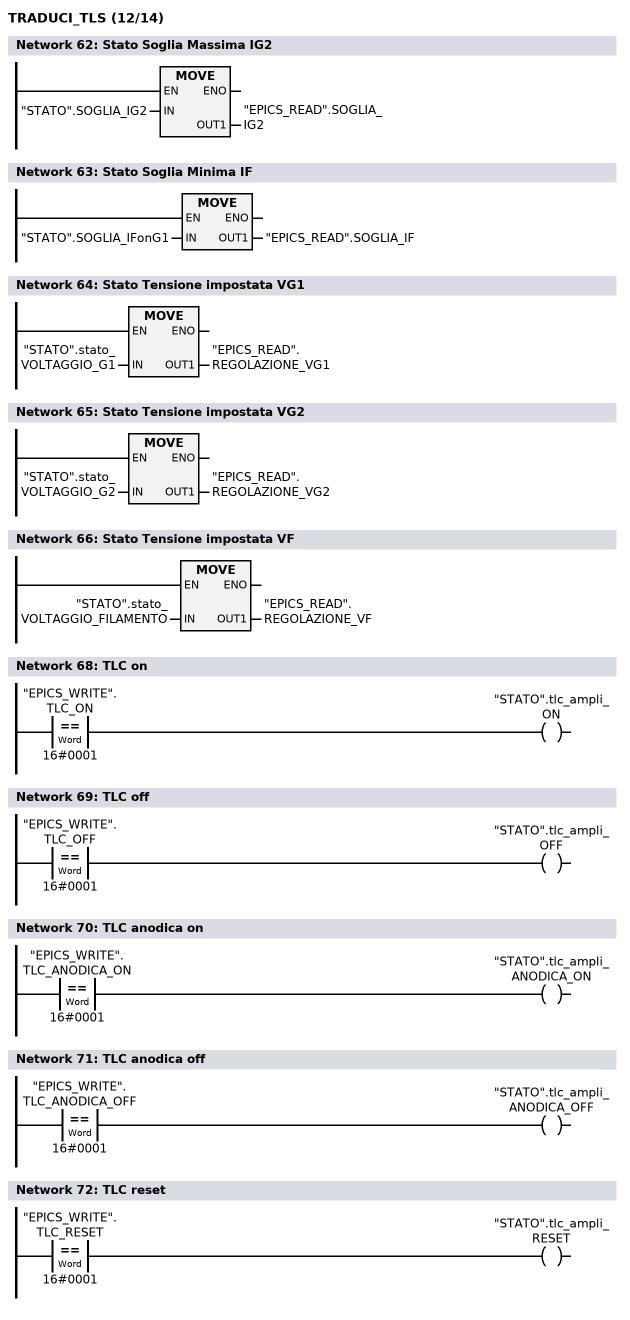
   RUNG wire#powerrail
      Move(in := "STATO".SOGLIA_IG2, out1 => "EPICS_READ".SOGLIA_IG2)
   END_RUNG
   // the same network as SCL:
   "EPICS_READ".SOGLIA_IG2 := "STATO".SOGLIA_IG2;
END_REGION

REGION Network 63: Stato Soglia Minima IF
   RUNG wire#powerrail
      Move(in := "STATO".SOGLIA_IFonG1, out1 => "EPICS_READ".SOGLIA_IF)
   END_RUNG
   // the same network as SCL:
   "EPICS_READ".SOGLIA_IF := "STATO".SOGLIA_IFonG1;
END_REGION

REGION Network 64: Stato Tensione impostata VG1
   RUNG wire#powerrail
      Move(in := "STATO".stato_VOLTAGGIO_G1, out1 => "EPICS_READ".REGOLAZIONE_VG1)
   END_RUNG
   // the same network as SCL:
   "EPICS_READ".REGOLAZIONE_VG1 := "STATO".stato_VOLTAGGIO_G1;
END_REGION

REGION Network 65: Stato Tensione impostata VG2
   RUNG wire#powerrail
      Move(in := "STATO".stato_VOLTAGGIO_G2, out1 => "EPICS_READ".REGOLAZIONE_VG2)
   END_RUNG
   // the same network as SCL:
   "EPICS_READ".REGOLAZIONE_VG2 := "STATO".stato_VOLTAGGIO_G2;
END_REGION

REGION Network 66: Stato Tensione impostata VF
   RUNG wire#powerrail
      Move(in := "STATO".stato_VOLTAGGIO_FILAMENTO, out1 => "EPICS_READ".REGOLAZIONE_VF)
   END_RUNG
   // the same network as SCL:
   "EPICS_READ".REGOLAZIONE_VF := "STATO".stato_VOLTAGGIO_FILAMENTO;
END_REGION

REGION Network 68: TLC on
   RUNG wire#powerrail
      { S7_Templates := "SrcType := Word" } EQ_Contact(in1 := "EPICS_WRITE".TLC_ON, in2 := 16#0001)
      Coil( "STATO".tlc_ampli_ON )
   END_RUNG
   // the same network as SCL:
   "STATO".tlc_ampli_ON := "EPICS_WRITE".TLC_ON = 16#0001;
END_REGION

REGION Network 69: TLC off
   RUNG wire#powerrail
      { S7_Templates := "SrcType := Word" } EQ_Contact(in1 := "EPICS_WRITE".TLC_OFF, in2 := 16#0001)
      Coil( "STATO".tlc_ampli_OFF )
   END_RUNG
   // the same network as SCL:
   "STATO".tlc_ampli_OFF := "EPICS_WRITE".TLC_OFF = 16#0001;
END_REGION

REGION Network 70: TLC anodica on
   RUNG wire#powerrail
      { S7_Templates := "SrcType := Word" } EQ_Contact(in1 := "EPICS_WRITE".TLC_ANODICA_ON, in2 := 16#0001)
      Coil( "STATO".tlc_ampli_ANODICA_ON )
   END_RUNG
   // the same network as SCL:
   "STATO".tlc_ampli_ANODICA_ON := "EPICS_WRITE".TLC_ANODICA_ON = 16#0001;
END_REGION

REGION Network 71: TLC anodica off
   RUNG wire#powerrail
      { S7_Templates := "SrcType := Word" } EQ_Contact(in1 := "EPICS_WRITE".TLC_ANODICA_OFF, in2 := 16#0001)
      Coil( "STATO".tlc_ampli_ANODICA_OFF )
   END_RUNG
   // the same network as SCL:
   "STATO".tlc_ampli_ANODICA_OFF := "EPICS_WRITE".TLC_ANODICA_OFF = 16#0001;
END_REGION

REGION Network 72: TLC reset
   RUNG wire#powerrail
      { S7_Templates := "SrcType := Word" } EQ_Contact(in1 := "EPICS_WRITE".TLC_RESET, in2 := 16#0001)
      Coil( "STATO".tlc_ampli_RESET )
   END_RUNG
   // the same network as SCL:
   "STATO".tlc_ampli_RESET := "EPICS_WRITE".TLC_RESET = 16#0001;
END_REGION

REGION Network 73: TLC imposta normal mode
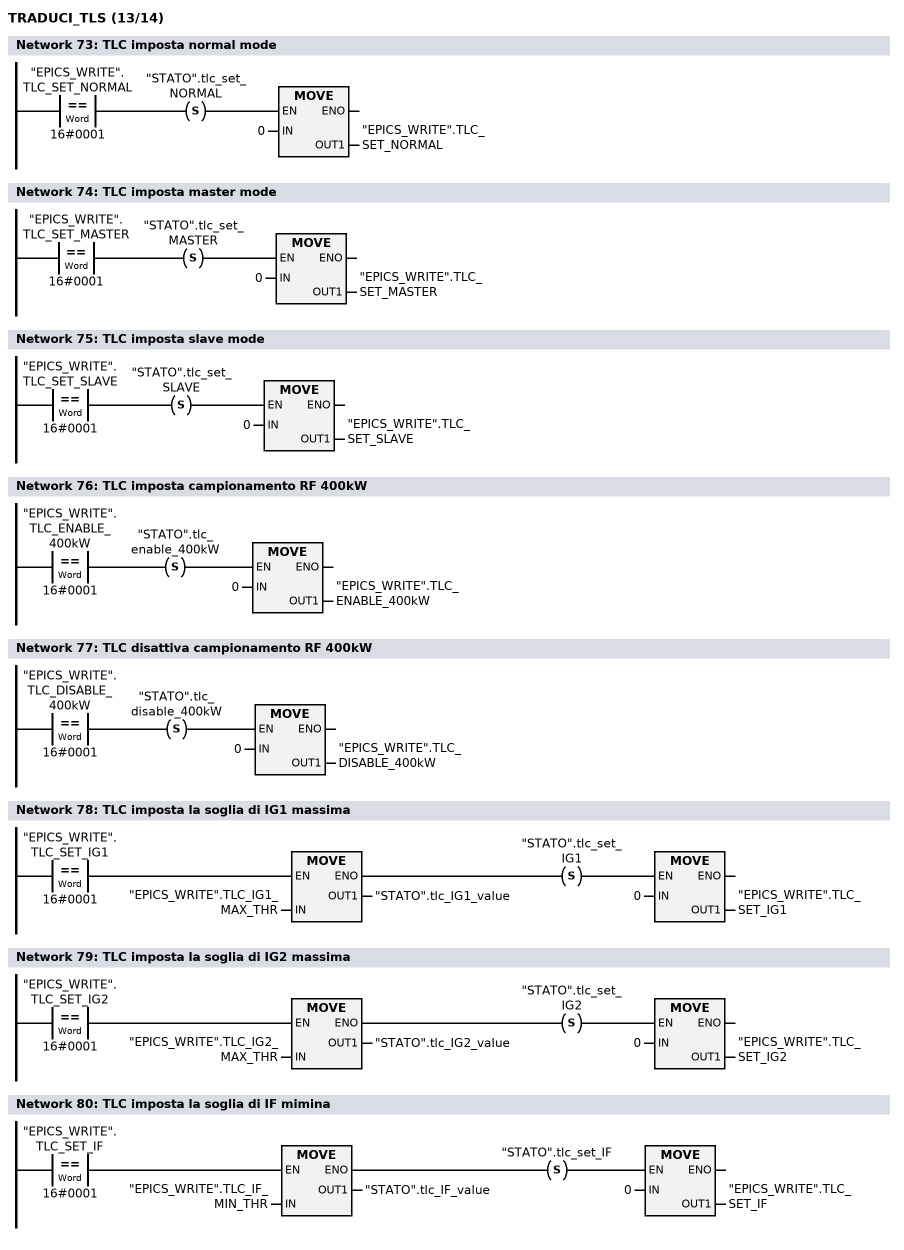
   RUNG wire#powerrail
      { S7_Templates := "SrcType := Word" } EQ_Contact(in1 := "EPICS_WRITE".TLC_SET_NORMAL, in2 := 16#0001)
      S_Coil( "STATO".tlc_set_NORMAL )
      Move(in := 0, out1 => "EPICS_WRITE".TLC_SET_NORMAL)
   END_RUNG
   // the same network as SCL:
   IF "EPICS_WRITE".TLC_SET_NORMAL = 16#0001 THEN
       "STATO".tlc_set_NORMAL := TRUE;
       "EPICS_WRITE".TLC_SET_NORMAL := 0;
   END_IF;
END_REGION

REGION Network 74: TLC imposta master mode
   RUNG wire#powerrail
      { S7_Templates := "SrcType := Word" } EQ_Contact(in1 := "EPICS_WRITE".TLC_SET_MASTER, in2 := 16#0001)
      S_Coil( "STATO".tlc_set_MASTER )
      Move(in := 0, out1 => "EPICS_WRITE".TLC_SET_MASTER)
   END_RUNG
   // the same network as SCL:
   IF "EPICS_WRITE".TLC_SET_MASTER = 16#0001 THEN
       "STATO".tlc_set_MASTER := TRUE;
       "EPICS_WRITE".TLC_SET_MASTER := 0;
   END_IF;
END_REGION

REGION Network 75: TLC imposta slave mode
   RUNG wire#powerrail
      { S7_Templates := "SrcType := Word" } EQ_Contact(in1 := "EPICS_WRITE".TLC_SET_SLAVE, in2 := 16#0001)
      S_Coil( "STATO".tlc_set_SLAVE )
      Move(in := 0, out1 => "EPICS_WRITE".TLC_SET_SLAVE)
   END_RUNG
   // the same network as SCL:
   IF "EPICS_WRITE".TLC_SET_SLAVE = 16#0001 THEN
       "STATO".tlc_set_SLAVE := TRUE;
       "EPICS_WRITE".TLC_SET_SLAVE := 0;
   END_IF;
END_REGION

REGION Network 76: TLC imposta campionamento RF 400kW
   RUNG wire#powerrail
      { S7_Templates := "SrcType := Word" } EQ_Contact(in1 := "EPICS_WRITE".TLC_ENABLE_400kW, in2 := 16#0001)
      S_Coil( "STATO".tlc_enable_400kW )
      Move(in := 0, out1 => "EPICS_WRITE".TLC_ENABLE_400kW)
   END_RUNG
   // the same network as SCL:
   IF "EPICS_WRITE".TLC_ENABLE_400kW = 16#0001 THEN
       "STATO".tlc_enable_400kW := TRUE;
       "EPICS_WRITE".TLC_ENABLE_400kW := 0;
   END_IF;
END_REGION

REGION Network 77: TLC disattiva campionamento RF 400kW
   RUNG wire#powerrail
      { S7_Templates := "SrcType := Word" } EQ_Contact(in1 := "EPICS_WRITE".TLC_DISABLE_400kW, in2 := 16#0001)
      S_Coil( "STATO".tlc_disable_400kW )
      Move(in := 0, out1 => "EPICS_WRITE".TLC_DISABLE_400kW)
   END_RUNG
   // the same network as SCL:
   IF "EPICS_WRITE".TLC_DISABLE_400kW = 16#0001 THEN
       "STATO".tlc_disable_400kW := TRUE;
       "EPICS_WRITE".TLC_DISABLE_400kW := 0;
   END_IF;
END_REGION

REGION Network 78: TLC imposta la soglia di IG1 massima
   RUNG wire#powerrail
      { S7_Templates := "SrcType := Word" } EQ_Contact(in1 := "EPICS_WRITE".TLC_SET_IG1, in2 := 16#0001)
      Move(in := "EPICS_WRITE".TLC_IG1_MAX_THR, out1 => "STATO".tlc_IG1_value)
      S_Coil( "STATO".tlc_set_IG1 )
      Move(in := 0, out1 => "EPICS_WRITE".TLC_SET_IG1)
   END_RUNG
   // the same network as SCL:
   IF "EPICS_WRITE".TLC_SET_IG1 = 16#0001 THEN
       "STATO".tlc_IG1_value := "EPICS_WRITE".TLC_IG1_MAX_THR;
       "STATO".tlc_set_IG1 := TRUE;
       "EPICS_WRITE".TLC_SET_IG1 := 0;
   END_IF;
END_REGION

REGION Network 79: TLC imposta la soglia di IG2 massima
   RUNG wire#powerrail
      { S7_Templates := "SrcType := Word" } EQ_Contact(in1 := "EPICS_WRITE".TLC_SET_IG2, in2 := 16#0001)
      Move(in := "EPICS_WRITE".TLC_IG2_MAX_THR, out1 => "STATO".tlc_IG2_value)
      S_Coil( "STATO".tlc_set_IG2 )
      Move(in := 0, out1 => "EPICS_WRITE".TLC_SET_IG2)
   END_RUNG
   // the same network as SCL:
   IF "EPICS_WRITE".TLC_SET_IG2 = 16#0001 THEN
       "STATO".tlc_IG2_value := "EPICS_WRITE".TLC_IG2_MAX_THR;
       "STATO".tlc_set_IG2 := TRUE;
       "EPICS_WRITE".TLC_SET_IG2 := 0;
   END_IF;
END_REGION

REGION Network 80: TLC imposta la soglia di IF mimina
   RUNG wire#powerrail
      { S7_Templates := "SrcType := Word" } EQ_Contact(in1 := "EPICS_WRITE".TLC_SET_IF, in2 := 16#0001)
      Move(in := "EPICS_WRITE".TLC_IF_MIN_THR, out1 => "STATO".tlc_IF_value)
      S_Coil( "STATO".tlc_set_IF )
      Move(in := 0, out1 => "EPICS_WRITE".TLC_SET_IF)
   END_RUNG
   // the same network as SCL:
   IF "EPICS_WRITE".TLC_SET_IF = 16#0001 THEN
       "STATO".tlc_IF_value := "EPICS_WRITE".TLC_IF_MIN_THR;
       "STATO".tlc_set_IF := TRUE;
       "EPICS_WRITE".TLC_SET_IF := 0;
   END_IF;
END_REGION

REGION Network 81: TLC imposta il DAC dell'anodica
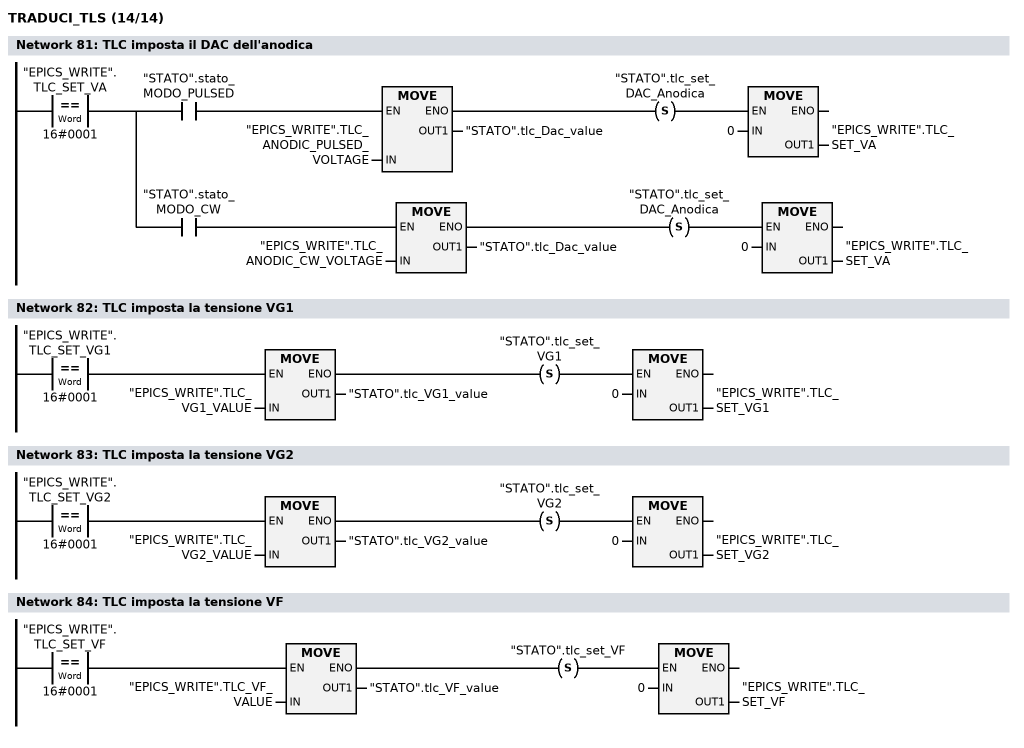
   RUNG wire#powerrail
      { S7_Templates := "SrcType := Word" } EQ_Contact(in1 := "EPICS_WRITE".TLC_SET_VA, in2 := 16#0001)
      wire#w1
      Contact( "STATO".stato_MODO_PULSED )
      Move(in := "EPICS_WRITE".TLC_ANODIC_PULSED_VOLTAGE, out1 => "STATO".tlc_Dac_value)
      S_Coil( "STATO".tlc_set_DAC_Anodica )
      Move(in := 0, out1 => "EPICS_WRITE".TLC_SET_VA)
   END_RUNG
   RUNG wire#w1
      Contact( "STATO".stato_MODO_CW )
      Move(in := "EPICS_WRITE".TLC_ANODIC_CW_VOLTAGE, out1 => "STATO".tlc_Dac_value)
      S_Coil( "STATO".tlc_set_DAC_Anodica )
      Move(in := 0, out1 => "EPICS_WRITE".TLC_SET_VA)
   END_RUNG
   // the same network as SCL:
   #_w1 := "EPICS_WRITE".TLC_SET_VA = 16#0001;
   IF #_w1 AND "STATO".stato_MODO_PULSED THEN
       "STATO".tlc_Dac_value := "EPICS_WRITE".TLC_ANODIC_PULSED_VOLTAGE;
       "STATO".tlc_set_DAC_Anodica := TRUE;
       "EPICS_WRITE".TLC_SET_VA := 0;
   END_IF;
   IF #_w1 AND "STATO".stato_MODO_CW THEN
       "STATO".tlc_Dac_value := "EPICS_WRITE".TLC_ANODIC_CW_VOLTAGE;
       "STATO".tlc_set_DAC_Anodica := TRUE;
       "EPICS_WRITE".TLC_SET_VA := 0;
   END_IF;
END_REGION

REGION Network 82: TLC imposta la tensione VG1
   RUNG wire#powerrail
      { S7_Templates := "SrcType := Word" } EQ_Contact(in1 := "EPICS_WRITE".TLC_SET_VG1, in2 := 16#0001)
      Move(in := "EPICS_WRITE".TLC_VG1_VALUE, out1 => "STATO".tlc_VG1_value)
      S_Coil( "STATO".tlc_set_VG1 )
      Move(in := 0, out1 => "EPICS_WRITE".TLC_SET_VG1)
   END_RUNG
   // the same network as SCL:
   IF "EPICS_WRITE".TLC_SET_VG1 = 16#0001 THEN
       "STATO".tlc_VG1_value := "EPICS_WRITE".TLC_VG1_VALUE;
       "STATO".tlc_set_VG1 := TRUE;
       "EPICS_WRITE".TLC_SET_VG1 := 0;
   END_IF;
END_REGION

REGION Network 83: TLC imposta la tensione VG2
   RUNG wire#powerrail
      { S7_Templates := "SrcType := Word" } EQ_Contact(in1 := "EPICS_WRITE".TLC_SET_VG2, in2 := 16#0001)
      Move(in := "EPICS_WRITE".TLC_VG2_VALUE, out1 => "STATO".tlc_VG2_value)
      S_Coil( "STATO".tlc_set_VG2 )
      Move(in := 0, out1 => "EPICS_WRITE".TLC_SET_VG2)
   END_RUNG
   // the same network as SCL:
   IF "EPICS_WRITE".TLC_SET_VG2 = 16#0001 THEN
       "STATO".tlc_VG2_value := "EPICS_WRITE".TLC_VG2_VALUE;
       "STATO".tlc_set_VG2 := TRUE;
       "EPICS_WRITE".TLC_SET_VG2 := 0;
   END_IF;
END_REGION

REGION Network 84: TLC imposta la tensione VF
   RUNG wire#powerrail
      { S7_Templates := "SrcType := Word" } EQ_Contact(in1 := "EPICS_WRITE".TLC_SET_VF, in2 := 16#0001)
      Move(in := "EPICS_WRITE".TLC_VF_VALUE, out1 => "STATO".tlc_VF_value)
      S_Coil( "STATO".tlc_set_VF )
      Move(in := 0, out1 => "EPICS_WRITE".TLC_SET_VF)
   END_RUNG
   // the same network as SCL:
   IF "EPICS_WRITE".TLC_SET_VF = 16#0001 THEN
       "STATO".tlc_VF_value := "EPICS_WRITE".TLC_VF_VALUE;
       "STATO".tlc_set_VF := TRUE;
       "EPICS_WRITE".TLC_SET_VF := 0;
   END_IF;
END_REGION
END_FUNCTION

FUNCTION "REGOLA_VG1" : Void   // FC13, LAD
{ S7_Optimized_Access := 'FALSE' }
VERSION : 0.1
BEGIN

REGION Network 1
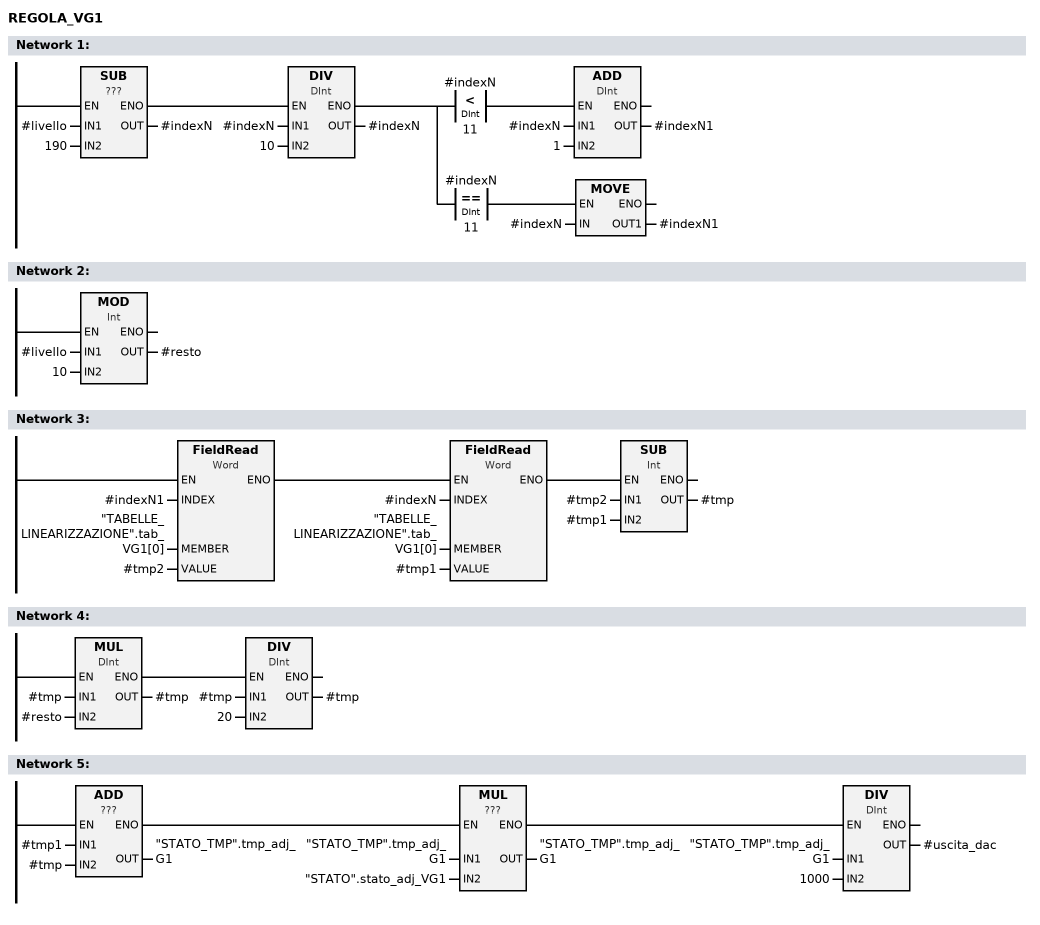
   RUNG wire#powerrail
      { S7_Templates := "SrcType := ???" } Sub(in1 := #livello, in2 := 190, out => #indexN)
      { S7_Templates := "SrcType := DInt" } Div(in1 := #indexN, in2 := 10, out => #indexN)
      wire#w1
      { S7_Templates := "SrcType := DInt" } LT_Contact(in1 := #indexN, in2 := 11)
      { S7_Templates := "SrcType := DInt" } Add(in1 := #indexN, in2 := 1, out => #indexN1)
   END_RUNG
   RUNG wire#w1
      { S7_Templates := "SrcType := DInt" } EQ_Contact(in1 := #indexN, in2 := 11)
      Move(in := #indexN, out1 => #indexN1)
   END_RUNG
   // the same network as SCL:
   #indexN := #livello - 190;
   #indexN := #indexN / 10;
   IF #indexN < 11 THEN #indexN1 := #indexN + 1; END_IF;
   IF #indexN = 11 THEN #indexN1 := #indexN; END_IF;
END_REGION

REGION Network 2
   RUNG wire#powerrail
      { S7_Templates := "SrcType := Int" } Mod(in1 := #livello, in2 := 10, out => #resto)
   END_RUNG
   // the same network as SCL:
   #resto := #livello MOD 10;
END_REGION

REGION Network 3
   // no SCL statement known for FieldRead: written as a call
   // ENO of a box is taken as its EN; it also drops when the box reports an error
   FieldRead(index := #indexN1, member := "TABELLE_LINEARIZZAZIONE".tab_VG1[0], value := #tmp2);
   FieldRead(index := #indexN, member := "TABELLE_LINEARIZZAZIONE".tab_VG1[0], value := #tmp1);
   #tmp := #tmp2 - #tmp1;
END_REGION

REGION Network 4
   RUNG wire#powerrail
      { S7_Templates := "SrcType := DInt" } Mul(in1 := #tmp, in2 := #resto, out => #tmp)
      { S7_Templates := "SrcType := DInt" } Div(in1 := #tmp, in2 := 20, out => #tmp)
   END_RUNG
   // the same network as SCL:
   #tmp := #tmp * #resto;
   #tmp := #tmp / 20;
END_REGION

REGION Network 5
   RUNG wire#powerrail
      { S7_Templates := "SrcType := ???" } Add(in1 := #tmp1, in2 := #tmp, out => "STATO_TMP".tmp_adj_G1)
      { S7_Templates := "SrcType := ???" } Mul(in1 := "STATO_TMP".tmp_adj_G1, in2 := "STATO".stato_adj_VG1, out => "STATO_TMP".tmp_adj_G1)
      { S7_Templates := "SrcType := DInt" } Div(in1 := "STATO_TMP".tmp_adj_G1, in2 := 1000, out => #uscita_dac)
   END_RUNG
   // the same network as SCL:
   "STATO_TMP".tmp_adj_G1 := #tmp1 + #tmp;
   "STATO_TMP".tmp_adj_G1 := "STATO_TMP".tmp_adj_G1 * "STATO".stato_adj_VG1;
   #uscita_dac := "STATO_TMP".tmp_adj_G1 / 1000;
END_REGION
END_FUNCTION

ORGANIZATION_BLOCK "Main"   // OB1, LAD, ProgramCycle
TITLE = "Main Program Sweep (Cycle)"
{ S7_Optimized_Access := 'FALSE' }
VERSION : 0.1
// ACCENSIONE LOGICA
BEGIN

REGION Network 1: Riconfiguro la porta di ricezione RS485
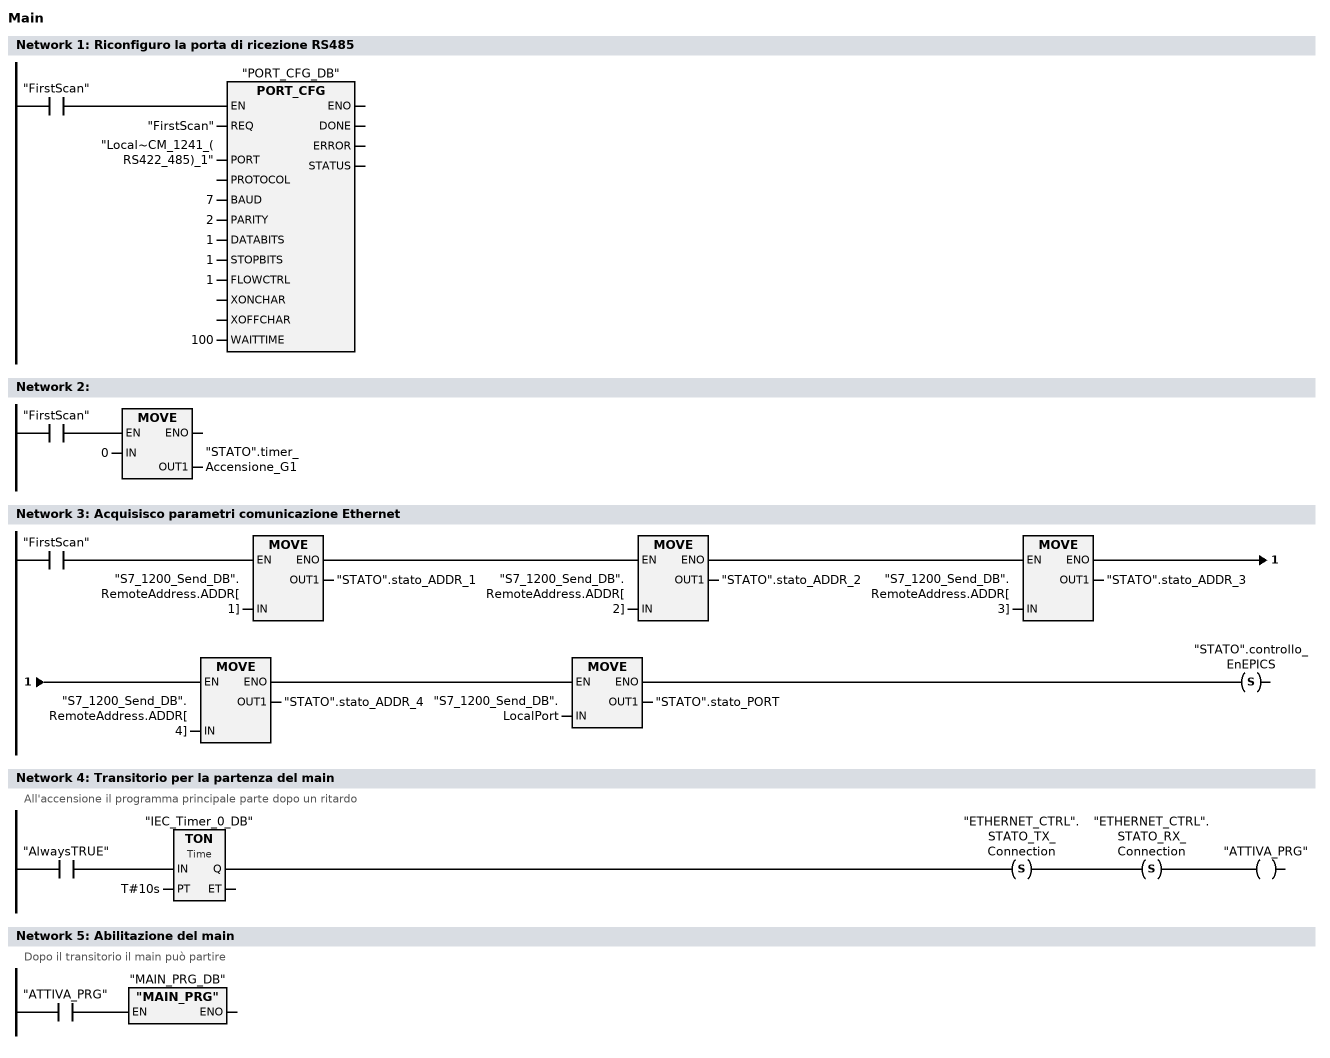
   IF "FirstScan" THEN
       "PORT_CFG_DB"(REQ := "FirstScan",   // PORT_CFG
                     PORT := "Local~CM_1241_(RS422_485)_1",
                     BAUD := 7,
                     PARITY := 2,
                     DATABITS := 1,
                     STOPBITS := 1,
                     FLOWCTRL := 1,
                     WAITTIME := 100);
   END_IF;
END_REGION

REGION Network 2
   RUNG wire#powerrail
      Contact( "FirstScan" )
      Move(in := 0, out1 => "STATO".timer_Accensione_G1)
   END_RUNG
   // the same network as SCL:
   IF "FirstScan" THEN "STATO".timer_Accensione_G1 := 0; END_IF;
END_REGION

REGION Network 3: Acquisisco parametri comunicazione Ethernet
   RUNG wire#powerrail
      Contact( "FirstScan" )
      Move(in := "S7_1200_Send_DB".RemoteAddress.ADDR[1], out1 => "STATO".stato_ADDR_1)
      Move(in := "S7_1200_Send_DB".RemoteAddress.ADDR[2], out1 => "STATO".stato_ADDR_2)
      Move(in := "S7_1200_Send_DB".RemoteAddress.ADDR[3], out1 => "STATO".stato_ADDR_3)
      Move(in := "S7_1200_Send_DB".RemoteAddress.ADDR[4], out1 => "STATO".stato_ADDR_4)
      Move(in := "S7_1200_Send_DB".LocalPort, out1 => "STATO".stato_PORT)
      S_Coil( "STATO".controllo_EnEPICS )
   END_RUNG
   // the same network as SCL:
   IF "FirstScan" THEN
       "STATO".stato_ADDR_1 := "S7_1200_Send_DB".RemoteAddress.ADDR[1];
       "STATO".stato_ADDR_2 := "S7_1200_Send_DB".RemoteAddress.ADDR[2];
       "STATO".stato_ADDR_3 := "S7_1200_Send_DB".RemoteAddress.ADDR[3];
       "STATO".stato_ADDR_4 := "S7_1200_Send_DB".RemoteAddress.ADDR[4];
       "STATO".stato_PORT := "S7_1200_Send_DB".LocalPort;
       "STATO".controllo_EnEPICS := TRUE;
   END_IF;
END_REGION

REGION Network 4: Transitorio per la partenza del main
   // All'accensione il programma principale parte dopo un ritardo
   "IEC_Timer_0_DB".TON(IN := "AlwaysTRUE", PT := T#10s);
   IF "IEC_Timer_0_DB".Q THEN
       "ETHERNET_CTRL".STATO_TX_Connection := TRUE;
       "ETHERNET_CTRL".STATO_RX_Connection := TRUE;
   END_IF;
   "ATTIVA_PRG" := "IEC_Timer_0_DB".Q;
END_REGION

REGION Network 5: Abilitazione del main
   // Dopo il transitorio il main può partire
   RUNG wire#powerrail
      Contact( "ATTIVA_PRG" )
      "MAIN_PRG_DB"()
   END_RUNG
   // the same network as SCL:
   IF "ATTIVA_PRG" THEN
       "MAIN_PRG_DB"();   // "MAIN_PRG"
   END_IF;
END_REGION
END_ORGANIZATION_BLOCK